(* Logix 5000 project; controller PLC_MCC1300_75F1 vendor 1 type 14 code 166 rev 32.11; software revision 32.04; part 61 of 83 *)
(* tags used below, declared in another part *)
   GP_ScadaPlate : GP_ScadaPlate;
   M311 : MAC_Conveyor;
   M315B : MAC_Conveyor;
   M315B_ALM : MAC_Conveyor_ALM;
   M315B_Data : UDT_Convoy_SL;
   M315B_HMR : MAC_Conveyor_HMR;
   M315B_HMW : MAC_Conveyor_HMW;
   M315B_SpaceConv_Utilities : SpaceConv_Utilities;
   M315Popup : MAC_Popup_ZC[2];
   M315Popup_ALM : MAC_Popup_ZC_ALM[2];
   M315Popup_HMR : MAC_Popup_ZC_HMR[2];
   M315Popup_HMW : MAC_Popup_ZC_HMW[2];
   O : INT[128];
   TMP_dHalfConveyorLength : DINT;
   TMP_xEnableZoneCleaning : BOOL;
   xAlwaysOFF : BOOL;
   xAlwaysON : BOOL;
   Z300_Conveyor : UDT_StandConv[29];
   Z300_LineTracking : UDT_LINE_TRACKING;
   Z301 : MAC_Zone_ML;
   Z402 : MAC_Zone;
   Z402_HMI_rgtPlateScada_Internal : HMI_LiteData[5,2,7];
(* MainProgram, continued *)

   // End load reentry (from M403) NEGATIVE
   50: XIC(M315B.PH_x.28)[GRT(M315B_SpaceConv_Utilities.O_dHeadPosition_cmm,M315B.AUX_dPresetStopLoad_cmm) XIO(M311.INPUT_xSyncroPhotocell_1) ,GRT(M315B_SpaceConv_Utilities.O_dHeadPosition_cmm,500000) ][OTE(M315B.PH_x.29) ,OTU(M315B.PH_x.28) ,NEQ(M315B_SpaceConv_Utilities.O_dHeadPosition_cmm,0) OTL(M315B.ST_xPlatePresence) ];
   // #####_HMI_STATUSES_#####
   51: NOP();
   // PhotocelPresence {x|x|x|x|O}
   52: XIC(M315B.INPUT_xSyncroPhotocell_1)OTE(M315B_HMR.xSensorPresence1);
   // PhotocelPresence {x|x|x|x|O}
   53: XIC(M315B.INPUT_xSyncroPhotocell_2)OTE(M315B_HMR.xSensorPresence2);
   // Manual Mode Enable {x|x|x|x|O}
   54: XIC(M315B.ST_xManualMode)OTE(M315B_HMR.xManualCommandEnabled);
   // Command forward M3
   55: XIC(M315B.ST_xManualMode)XIC(M315B_HMW.rgxMan.4)XIC(M315B.OUTPUT_xRun_M1)OTE(M315B_HMR.rgxMan.4);
   // Command backward M3
   56: XIC(M315B.ST_xManualMode)XIC(M315B_HMW.rgxMan.5)XIC(M315B.OUTPUT_xReverse_M1)OTE(M315B_HMR.rgxMan.5);
   // Command forward M4
   57: XIC(M315B.ST_xManualMode)XIC(M315B_HMW.rgxMan.6)XIC(M315B.OUTPUT_xRun_M2)OTE(M315B_HMR.rgxMan.6);
   // Command backward M4
   58: XIC(M315B.ST_xManualMode)XIC(M315B_HMW.rgxMan.7)XIC(M315B.OUTPUT_xReverse_M2)OTE(M315B_HMR.rgxMan.7);
   // Cleaning Enabled {x|x|x|x|O}
   59: XIC(M315B.ST_xCleaningAccepted)[XIC(Z402.ST_xCleaningAccepted) ,XIO(TMP_xEnableZoneCleaning) ]OTE(M315B_HMR.xCleaningEnabled);
   // Virtual door Enabled {x|x|x|x|O}
   60: XIC(M315B.ST_xVirtualDoorEnabled)OTE(M315B_HMR.xVirtualDoorEnabled);
   // Id plate presence
   61: XIC(M315B.ST_xIdPlatePresence)OTE(M315B_HMR.xIdPlatePresence);
   // Machine state M3
   62: XIC(xAlwaysON)[MOV(1,M315B_HMR.dState3) ,XIC(M315B.OUTPUT_xRun_M1) MOV(3,M315B_HMR.dState3) ,XIC(M315B.OUTPUT_xReverse_M1) MOV(4,M315B_HMR.dState3) ,XIC(M315B.ST_xMachineWarning) MOV(5,M315B_HMR.dState3) ,XIC(M315B.ST_xMachineAlarm) MOV(7,M315B_HMR.dState3) ];
   // Machine state M4
   63: XIC(xAlwaysON)[MOV(1,M315B_HMR.dState4) ,XIC(M315B.OUTPUT_xRun_M2) MOV(3,M315B_HMR.dState4) ,XIC(M315B.OUTPUT_xReverse_M2) MOV(4,M315B_HMR.dState4) ,XIC(M315B.ST_xMachineAlarm) MOV(7,M315B_HMR.dState4) ];
   // State Sensor
   64: XIC(xAlwaysON)[MOV(1,M315B_HMR.dStateSensor1) ,XIC(M315B_ALM.rgxWarning[0].0) MOV(7,M315B_HMR.dStateSensor1) ];
   // State Sensor
   65: XIC(xAlwaysON)[MOV(1,M315B_HMR.dStateSensor2) ,XIC(M315B_ALM.rgxWarning[0].1) MOV(7,M315B_HMR.dStateSensor2) ];
   66: XIC(M315B.ST_xIdPlatePresence)GP_ScadaPlate(GP_ScadaPlate,M315B_Data,0,M315B_SpaceConv_Utilities.O_dHeadPosition_cmm,M315B_SpaceConv_Utilities.CONST_dConveyorWidth_cmm,M315B_SpaceConv_Utilities.CONST_dConveyorLength_cmm,M315B_SpaceConv_Utilities.ST_xLastModLoadBkw,M315B_SpaceConv_Utilities.ST_xLastModUnloadBkw,1,0,Z402_HMI_rgtPlateScada_Internal);
END_ROUTINE

ROUTINE M315Popup0_Faults   (* ladder *)
   // Reset faults
   0: XIC(Z301.ST_xAlarmOff)FLL(0,M315Popup_ALM[0],1);
   1: XIC(Z300_Conveyor[27].ST_xOutputEnable)XIO(Z300_Conveyor[27].ST_xCleaningEnabled)XIC(M315Popup[0].ST_xEnableControlError)[[XIC(M315Popup[0].OUTPUT_xPopupLifting) XIO(M315Popup[0].INPUT_xPopupHigh) ,XIC(M315Popup[0].OUTPUT_xPopupDescent) XIO(M315Popup[0].INPUT_xPopupLow) ,XIO(M315Popup[0].INPUT_xPopupHigh) XIO(M315Popup[0].INPUT_xPopupLow) XIO(M315Popup_ALM[0].rgxStoppingFault[0].0) ] TON(M315Popup[0].tmON_LiftingTimeOut,?,?) ,[XIC(M315Popup[0].tmON_LiftingTimeOut.DN) ,XIC(M315Popup[0].INPUT_xPopupHigh) XIC(M315Popup[0].INPUT_xPopupLow) ] OTL(M315Popup_ALM[0].rgxStoppingFault[0].0) ];
   2: XIC(M315Popup[0].ST_xEnableControlError)XIO(M315Popup[0].INPUT_xLiftingProtectionMotor)OTL(M315Popup_ALM[0].rgxFault[0].0);
   3: XIC(M315Popup[0].ST_xEnableControlError)XIC(M315Popup[0].ST_xOutputEnable)[[XIC(M315Popup[0].OUTPUT_xPopupLifting) ,XIC(M315Popup[0].OUTPUT_xPopupDescent) ] XIO(M315Popup[0].INPUT_xLiftingFeedbackMotor) ,XIO(M315Popup[0].OUTPUT_xPopupLifting) XIO(M315Popup[0].OUTPUT_xPopupDescent) XIC(M315Popup[0].INPUT_xLiftingFeedbackMotor) ][TON(M315Popup[0].tmON_LiftingFeedbackTimeOut,?,?) ,XIC(M315Popup[0].tmON_LiftingFeedbackTimeOut.DN) OTL(M315Popup_ALM[0].rgxFault[0].1) ];
   4: XIC(M315Popup[0].ST_xEnableControlError)XIO(M315Popup[0].INPUT_xLiftingSafetySwitch)XIC(xAlwaysOFF)OTL(M315Popup_ALM[0].rgxFault[0].2);
   5: XIC(M315Popup[0].ST_xEnableControlError)XIO(M315Popup[0].INPUT_xProtectionCoolingFan)OTL(M315Popup_ALM[0].rgxFault[0].3);
   6: XIC(M315Popup[0].ST_xEnableControlError)XIO(M315Popup[0].INPUT_xFeedbackCoolingFan)OTL(M315Popup_ALM[0].rgxFault[0].4);
   // Stopped machine fault
   7: [NEQ(M315Popup_ALM[0].rgxStoppingFault[0],0) ,NEQ(M315Popup_ALM[0].rgxStoppingFault_M[0],0) ]OTE(M315Popup[0].ST_xStopMachineFault);
   // Stopped next cycle fault
   8: [NEQ(M315Popup_ALM[0].rgxFault[0],0) ,NEQ(M315Popup_ALM[0].rgxFault_M[0],0) ]OTE(M315Popup[0].ST_xStopNextCycleFault);
   9: XIC(M315Popup[0].ST_xEnableControlError)XIC(M315Popup[0].ST_xOutputEnable)[XIC(M315Popup[0].PH_xRise) XIO(M315Popup[0].ST_xInitialConditionForRise) XIO(M315Popup[0].INPUT_xPopupHigh) ,XIC(M315Popup[0].PH_xDescend) XIO(M315Popup[0].ST_xInitialConditionForDescend) XIO(M315Popup[0].INPUT_xPopupLow) ]OTE(M315Popup[0].ST_xMachineWarning);
END_ROUTINE

ROUTINE M315Popup0_Logic   (* ladder *)
   // #####_CONSTANTS_#####
   0: NOP();
   1: XIC(xAlwaysON)OTE(M315Popup[0].ST_xTunnelType);
   2: DIV(Z300_LineTracking.rgtTrkConv[27].dLengthConveyor,2,TMP_dHalfConveyorLength);
   3: MOV(Z300_LineTracking.rgtTrkConv[27].dStartPosition_cmm,M315Popup[0].AUX_dStartPosition_cmm)MOV(Z300_LineTracking.rgtTrkConv[27].dEndPosition_cmm,M315Popup[0].AUX_dEndPosition_cmm)MOV(1500,M315Popup[0].AUX_dReactionTime_ms)MOV(200000,M315Popup[0].AUX_dWindowSearch_cmm)MOV(Z300_Conveyor[27].AUX_rgdCurrentSpeed_mm_min[0],M315Popup[0].AUX_dSpeedConveyor_mm_min);
   // #####_MATCH_#####
   4: NOP();
   5: XIC(Z301.ST_xEnableControlError)OTE(M315Popup[0].ST_xEnableControlError);
   // #####_ALARMS_#####
   6: NOP();
   7: JSR(M315Popup0_Faults,0);
   // #####_HMI_LOGICS_#####
   8: NOP();
   9: XIC(xAlwaysON)OTE(M315Popup[0].ST_xExternalConditionToRise);
   // #####_STATUSES_#####
   10: NOP();
   11: [XIC(M315Popup[0].ST_xStopMachineFault) ,XIC(M315Popup[0].ST_xStopNextCycleFault) ]OTE(M315Popup[0].ST_xMachineAlarm);
   12: [XIO(M315Popup[0].ST_xPhasesInProgress) ,XIO(M315Popup[0].ST_xOutputEnable) ]OTE(M315Popup[0].ST_xConditionOKForStopCycle);
   13: XIC(Z301.ST_xCycleON)XIO(M315Popup[0].ST_xManualMode)XIO(M315Popup[0].ST_xMachineAlarm)OTE(M315Popup[0].ST_xOutputEnable);
   14: XIC(Z301.ST_xCycleON)XIC(M315Popup[0].ST_xOutputEnable)XIO(M315Popup[0].ST_xPhasesInProgress)XIO(M315Popup[0].INPUT_xPopupHigh)XIC(M315Popup[0].INPUT_xPopupLow)XIO(M315Popup[0].ST_xCleaningAccepted)OTE(M315Popup[0].ST_xInitialConditionForRise);
   15: XIC(Z301.ST_xCycleON)XIC(M315Popup[0].ST_xOutputEnable)XIO(M315Popup[0].ST_xPhasesInProgress)XIO(M315Popup[0].INPUT_xPopupLow)XIC(M315Popup[0].INPUT_xPopupHigh)XIO(M315Popup[0].ST_xCleaningAccepted)OTE(M315Popup[0].ST_xInitialConditionForDescend);
   16: [XIC(M315Popup_HMW[0].xEnableDisableManualCommand) XIC(xAlwaysOFF) ,XIC(Z300_Conveyor[27].ST_xManualCmdEnabled) ]XIC(M315Popup[0].ST_xConditionOKForStopCycle)XIC(M315Popup[1].ST_xConditionOKForStopCycle)OTE(M315Popup[0].ST_xManualMode);
   17: XIO(M315Popup[0].ST_xManualMode)MOV(0,M315Popup_HMW[0].rgxMan);
   // #####_PHASES_&_LOGICS_#####
   18: NOP();
   19: XIC(xAlwaysON)OTE(M315Popup[0].ST_xCleaningConditionOK);
   20: [XIC(M315Popup_HMW[0].xLocalCleaningRequest) XIC(xAlwaysOFF) ,XIC(Z300_Conveyor[27].ST_xCleaningEnabled) XIC(M315Popup[0].INPUT_xPopupLow) ][XIC(M315Popup[0].ST_xCleaningConditionOK) ,XIC(M315Popup[0].ST_xCleaningAccepted) ]OTE(M315Popup[0].ST_xCleaningAccepted);
   21: XIC(M315Popup[0].ST_xInitialConditionForRise)XIC(M315Popup[0].ST_xExternalConditionToRise)XIC(M315Popup[0].ST_xRequestRise)XIO(M315Popup[0].PH_xRise)OTL(M315Popup[0].PH_xRise);
   22: XIC(M315Popup[0].PH_xRise)XIC(M315Popup[0].INPUT_xPopupHigh)XIO(M315Popup[0].INPUT_xPopupLow)[OTU(M315Popup[0].PH_xRise) ,OTE(M315Popup[0].PH_xEndRise) ];
   23: XIC(M315Popup[0].ST_xInitialConditionForDescend)XIC(M315Popup[0].ST_xExternalConditionToDescend)XIC(M315Popup[0].ST_xRequestDescend)[XIC(M315Popup[1].ST_xRequestDescend) ,XIC(M315Popup[1].INPUT_xPopupLow) ]XIO(M315Popup[0].PH_xDescend)OTL(M315Popup[0].PH_xDescend);
   24: XIC(M315Popup[0].PH_xDescend)XIC(M315Popup[0].INPUT_xPopupLow)XIO(M315Popup[0].INPUT_xPopupHigh)[OTU(M315Popup[0].PH_xDescend) ,OTE(M315Popup[0].PH_xEndDescend) ];
   25: [XIC(M315Popup[0].PH_xRise) ,XIC(M315Popup[0].PH_xEndRise) ,XIC(M315Popup[0].PH_xDescend) ,XIC(M315Popup[0].PH_xEndDescend) ]OTE(M315Popup[0].ST_xPhasesInProgress);
   26: [XIC(M315Popup[0].PH_xEndDescend) ,XIO(xAlwaysOFF) XIC(M315Popup[0].INPUT_xPopupLow) ]OTU(M315Popup[0].ST_xPlatePresence);
   27: XIO(M315Popup[0].ST_xPhasesInProgress)[XIC(M315Popup[0].INPUT_xPopupLow) XIO(M315Popup[0].INPUT_xPopupHigh) ,XIC(M315Popup[0].ST_xTunnelType) XIC(M315Popup[0].INPUT_xPopupHigh) XIO(M315Popup[0].INPUT_xPopupLow) ]OTE(M315Popup[0].ST_xOutOfEncumbrance);
   28: XIO(M315Popup[0].ST_xPhasesInProgress)XIO(M315Popup[0].ST_xPlatePresence)XIO(M315Popup[0].INPUT_xPopupHigh)XIC(M315Popup[0].INPUT_xPopupLow)OTE(M315Popup[0].ST_xConditionToReceiveGlass);
   29: XIO(M315Popup[0].ST_xPhasesInProgress)XIC(M315Popup[0].INPUT_xPopupHigh)XIO(M315Popup[0].INPUT_xPopupLow)OTE(M315Popup[0].ST_xConditionForUpperConveyor);
   // #####_EXTERNAL_DEVICE_#####
   30: NOP();
   // #####_HMI_STATUSES_#####
   31: NOP();
   32: XIC(M315Popup[0].INPUT_xPopupHigh)OTE(M315Popup_HMR[0].xHighPosition);
   33: XIC(M315Popup[0].INPUT_xPopupLow)OTE(M315Popup_HMR[0].xLowPosition);
   34: [MOV(1,M315Popup_HMR[0].rgdState) ,[XIC(M315Popup[0].OUTPUT_xPopupLifting) ,XIC(M315Popup[0].OUTPUT_xPopupDescent) ] MOV(3,M315Popup_HMR[0].rgdState) ,XIC(M315Popup[0].ST_xMachineWarning) MOV(5,M315Popup_HMR[0].rgdState) ,XIC(M315Popup[0].ST_xMachineAlarm) MOV(7,M315Popup_HMR[0].rgdState) ];
   35: XIC(M315Popup[0].ST_xCleaningAccepted)OTE(M315Popup_HMR[0].xPopUpCleaningEnabled);
   36: XIC(M315Popup[0].ST_xManualMode)XIC(M315Popup_HMW[0].rgxMan.0)XIC(M315Popup[0].OUTPUT_xPopupLifting)OTE(M315Popup_HMR[0].rgxMan.0);
   37: XIC(M315Popup[0].ST_xManualMode)XIC(M315Popup_HMW[0].rgxMan.1)XIC(M315Popup[0].OUTPUT_xPopupDescent)OTE(M315Popup_HMR[0].rgxMan.1);
   38: XIC(M315Popup[0].ST_xManualMode)XIC(M315Popup_HMW[0].rgxMan.8)XIC(M315Popup[0].OUTPUT_xRun)OTE(M315Popup_HMR[0].rgxMan.8);
   39: XIC(M315Popup[0].ST_xManualMode)XIC(M315Popup_HMW[0].rgxMan.9)XIC(M315Popup[0].OUTPUT_xReverse)OTE(M315Popup_HMR[0].rgxMan.9);
END_ROUTINE

ROUTINE M315Popup1_Faults   (* ladder *)
   // Reset faults
   0: XIC(Z301.ST_xAlarmOff)FLL(0,M315Popup_ALM[1],1);
   1: XIC(Z300_Conveyor[28].ST_xOutputEnable)XIO(Z300_Conveyor[28].ST_xCleaningEnabled)XIC(M315Popup[1].ST_xEnableControlError)[[XIC(M315Popup[1].OUTPUT_xPopupLifting) XIO(M315Popup[1].INPUT_xPopupHigh) ,XIC(M315Popup[1].OUTPUT_xPopupDescent) XIO(M315Popup[1].INPUT_xPopupLow) ,XIO(M315Popup[1].INPUT_xPopupHigh) XIO(M315Popup[1].INPUT_xPopupLow) XIO(M315Popup_ALM[0].rgxStoppingFault[0].0) ] TON(M315Popup[1].tmON_LiftingTimeOut,?,?) ,[XIC(M315Popup[1].tmON_LiftingTimeOut.DN) ,XIC(M315Popup[1].INPUT_xPopupHigh) XIC(M315Popup[1].INPUT_xPopupLow) ] OTL(M315Popup_ALM[1].rgxStoppingFault[0].0) ];
   2: XIC(M315Popup[1].ST_xEnableControlError)XIO(M315Popup[1].INPUT_xLiftingProtectionMotor)OTL(M315Popup_ALM[1].rgxFault[0].0);
   3: XIC(M315Popup[1].ST_xEnableControlError)XIC(M315Popup[1].ST_xOutputEnable)[[XIC(M315Popup[1].OUTPUT_xPopupLifting) ,XIC(M315Popup[1].OUTPUT_xPopupDescent) ] XIO(M315Popup[1].INPUT_xLiftingFeedbackMotor) ,XIO(M315Popup[1].OUTPUT_xPopupLifting) XIO(M315Popup[1].OUTPUT_xPopupDescent) XIC(M315Popup[1].INPUT_xLiftingFeedbackMotor) ][TON(M315Popup[1].tmON_LiftingFeedbackTimeOut,?,?) ,XIC(M315Popup[1].tmON_LiftingFeedbackTimeOut.DN) OTL(M315Popup_ALM[1].rgxFault[0].1) ];
   4: XIC(M315Popup[1].ST_xEnableControlError)XIO(M315Popup[1].INPUT_xLiftingSafetySwitch)XIC(xAlwaysOFF)OTL(M315Popup_ALM[1].rgxFault[0].2);
   5: XIC(M315Popup[1].ST_xEnableControlError)XIO(M315Popup[1].INPUT_xProtectionCoolingFan)OTL(M315Popup_ALM[1].rgxFault[0].3);
   6: XIC(M315Popup[1].ST_xEnableControlError)XIO(M315Popup[1].INPUT_xFeedbackCoolingFan)OTL(M315Popup_ALM[1].rgxFault[0].4);
   // Stopped machine fault
   7: [NEQ(M315Popup_ALM[1].rgxStoppingFault[0],0) ,NEQ(M315Popup_ALM[1].rgxStoppingFault_M[0],0) ]OTE(M315Popup[1].ST_xStopMachineFault);
   // Stopped next cycle fault
   8: [NEQ(M315Popup_ALM[1].rgxFault[0],0) ,NEQ(M315Popup_ALM[1].rgxFault_M[0],0) ]OTE(M315Popup[1].ST_xStopNextCycleFault);
   9: XIC(M315Popup[1].ST_xEnableControlError)XIC(M315Popup[1].ST_xOutputEnable)[XIC(M315Popup[1].PH_xRise) XIO(M315Popup[1].ST_xInitialConditionForRise) XIO(M315Popup[1].INPUT_xPopupHigh) ,XIC(M315Popup[1].PH_xDescend) XIO(M315Popup[1].ST_xInitialConditionForDescend) XIO(M315Popup[1].INPUT_xPopupLow) ]OTE(M315Popup[1].ST_xMachineWarning);
END_ROUTINE
